// TIA Portal project "Lift" (V15.1)

(* hardware
DEVICE "S7-1200 station_1"  S7-1200 Station
   slot 0: "Rack_0"  S7-1200 Rack  Rack  V1.0
   slot 1: "PLC_1"  CPU 1215C DC/DC/DC  6ES7 215-1AG40-0XB0  V4.2
DEVICE "HMI_1"  TP1500 Basic color PN
   slot 0: "HMI_1"  TP1500 Basic color PN  6AV6 647-0AG11-3AX0  12.0.0.0
   slot 1: "HMI_RT_1"  TP1500 Basic color PN  6AV6 647-0AG11-3AX0  12.0.0.0
   slot 5: "HMI_1.IE_CP_1"  PROFINET Interface  12.0.0.0
      slot 1: "PROFINET Interface_1"  PROFINET Interface
         slot 1: "Port_1"  Port
DEVICE "HMI_2"  KTP700 Basic PN
   slot 0: "HMI_2"  KTP700 Basic PN  6AV2 123-2GB03-0AX0  15.1.0.0
   slot 1: "HMI_RT_2"  KTP700 Basic PN  6AV2 123-2GB03-0AX0  15.1.0.0
   slot 5: "HMI_2.IE_CP_1"  PROFINET Interface  15.0.1.0
      slot 1: "PROFINET Interface_1"  PROFINET Interface
         slot 1: "Port_1"  Port
*)

// ===== PLC "PLC_1"  CPU 1215C DC/DC/DC =====

VAR_GLOBAL   // PLC tag table "Default tag table"
   "Clock_Byte" AT %MB1 : Byte;
   "Clock_10Hz" AT %M1.0 : Bool;
   "Clock_5Hz" AT %M1.1 : Bool;
   "Clock_2.5Hz" AT %M1.2 : Bool;
   "Clock_2Hz" AT %M1.3 : Bool;
   "Clock_1.25Hz" AT %M1.4 : Bool;
   "Clock_1Hz" AT %M1.5 : Bool;
   "Clock_0.625Hz" AT %M1.6 : Bool;
   "Clock_0.5Hz" AT %M1.7 : Bool;
END_VAR

VAR_GLOBAL   // PLC tag table "lift butoane interior"
   "buton_parter" AT %I0.0 : Bool;
   "buton_et1" AT %I0.1 : Bool;
   "buton_et2" AT %I0.2 : Bool;
   "butor_urgenta" AT %I0.3 : Bool;
   "reset_button_urgenta" AT %I0.4 : Bool;
END_VAR

VAR_GLOBAL   // PLC tag table "lift outputs"
   "usa_parter" AT %Q0.0 : Bool;
   "usa_et1" AT %Q0.1 : Bool;
   "usa_et2" AT %Q0.2 : Bool;
   "bec_lift" AT %Q0.3 : Bool;
   "usa lift" AT %Q0.4 : Bool;
END_VAR

VAR_GLOBAL   // PLC tag table "lift auxiliares"
   "block_request_parter" AT %M0.0 : Bool;
   "urgenta_pressed" AT %M2.0 : Bool;
   "block_request_et1" AT %M2.1 : Bool;
   "block_request_et2" AT %M2.2 : Bool;
   "directie sus" AT %M2.3 : Bool;
   "directie jos" AT %M2.4 : Bool;
   "block_persoana" AT %M2.5 : Bool;
   "limitator_parter" AT %M2.6 : Bool;
   "limitator_1" AT %M2.7 : Bool;
   "limitator_2" AT %M3.0 : Bool;
   "reset_block_requests" AT %M3.1 : Bool;
   "tag_auxiliar_hmi" AT %M3.2 : Bool;
END_VAR

VAR_GLOBAL   // PLC tag table "lift butoane exterior"
   "buton_exterior_parter" AT %I0.5 : Bool;
   "buton_et1_ext" AT %I0.6 : Bool;
   "buton_et2_ext" AT %I0.7 : Bool;
END_VAR

VAR_GLOBAL   // PLC tag table "lift inputs(usi)"
   "usa_parter_i" AT %I1.0 : Bool;
   "usa_et1_i" AT %I1.1 : Bool;
   "usa_et2_i" AT %I1.2 : Bool;
   "usa_lift_i" AT %I1.3 : Bool;
END_VAR

DATA_BLOCK "motor_DB"   // DB1
{ S7_Optimized_Access := 'TRUE' }
VERSION : 0.1
// stored: InstanceOfName motor parter
"motor parter"
BEGIN
END_DATA_BLOCK

DATA_BLOCK "motor_DB_1"   // DB2
{ S7_Optimized_Access := 'TRUE' }
VERSION : 0.1
// stored: InstanceOfName motor parter
"motor parter"
BEGIN
END_DATA_BLOCK

DATA_BLOCK "motor_DB_2"   // DB3
{ S7_Optimized_Access := 'TRUE' }
VERSION : 0.1
// stored: InstanceOfName motor parter
"motor parter"
BEGIN
END_DATA_BLOCK

DATA_BLOCK "motor et1_DB"   // DB4
{ S7_Optimized_Access := 'TRUE' }
VERSION : 0.1
// stored: InstanceOfName motor et1
"motor et1"
BEGIN
END_DATA_BLOCK

DATA_BLOCK "motor et2_DB"   // DB5
{ S7_Optimized_Access := 'TRUE' }
VERSION : 0.1
// stored: InstanceOfName motor et2
"motor et2"
BEGIN
END_DATA_BLOCK

DATA_BLOCK "motor parter_DB"   // DB6
{ S7_Optimized_Access := 'TRUE' }
VERSION : 0.1
// stored: InstanceOfName motor parter
"motor parter"
BEGIN
END_DATA_BLOCK

DATA_BLOCK "motor et1_DB_1"   // DB7
{ S7_Optimized_Access := 'TRUE' }
VERSION : 0.1
// stored: InstanceOfName motor et1
"motor et1"
BEGIN
END_DATA_BLOCK

DATA_BLOCK "motor et2_DB_1"   // DB8
{ S7_Optimized_Access := 'TRUE' }
VERSION : 0.1
// stored: InstanceOfName motor et2
"motor et2"
BEGIN
END_DATA_BLOCK

DATA_BLOCK "Commands"   // DB9
{ S7_Optimized_Access := 'TRUE' }
VERSION : 0.1
   VAR
      buton_et1_ext : Bool;
      buton_et2_ext : Bool;
      buton_parter_ext : Bool;
      buton_et1_int : Bool;
      _buton_et2_int : Bool;
      buton_parter_int : Bool;
      buton_urgenta : Bool;
      buton_urgenta_reset : Bool;
      usa_lift_input : Bool;
   END_VAR
BEGIN
END_DATA_BLOCK

FUNCTION_BLOCK "motor parter"   // FB1, LAD
{ S7_Optimized_Access := 'TRUE' }
VERSION : 0.1
   VAR_INPUT
      req_p : Bool;
      et_p : Bool;
      et_1 : Bool;
      et_2 : Bool;
   END_VAR
   VAR_OUTPUT
      dir_sus : Bool;
      dir_jos : Bool;
   END_VAR
BEGIN

REGION Network 1: cerere de la parter
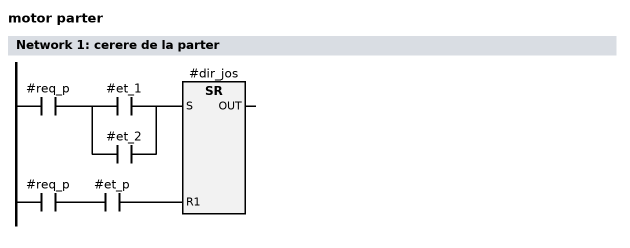
   RUNG wire#powerrail
      Contact( #req_p )
      wire#w1
      Contact( #et_1 )
      wire#w2
      S_SR(operand := #dir_jos, r1 := wire#w3)
   END_RUNG
   RUNG wire#w1
      Contact( #et_2 )
   END_RUNG wire#w2
   RUNG wire#powerrail
      Contact( #req_p )
      Contact( #et_p )
   END_RUNG wire#w3
   // the same network as SCL:
   IF #req_p AND (#et_1 OR #et_2) THEN
       #dir_jos := TRUE;   // SR flip-flop
   END_IF;
   IF #req_p AND #et_p THEN #dir_jos := FALSE; END_IF;
END_REGION
END_FUNCTION_BLOCK

FUNCTION_BLOCK "motor et2"   // FB2, LAD
{ S7_Optimized_Access := 'TRUE' }
VERSION : 0.1
   VAR_INPUT
      req_2 : Bool;
      et_p : Bool;
      et_1 : Bool;
      et_2 : Bool;
   END_VAR
   VAR_OUTPUT
      dir_sus : Bool;
      dir_jos : Bool;
   END_VAR
BEGIN

REGION Network 1: cerere de la etaj 2
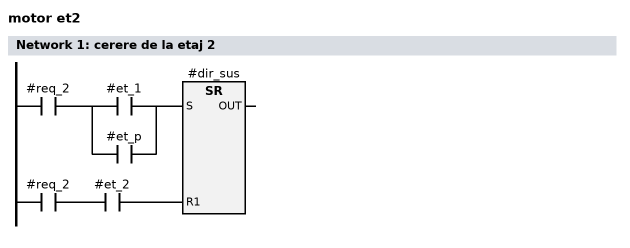
   RUNG wire#powerrail
      Contact( #req_2 )
      wire#w1
      Contact( #et_1 )
      wire#w2
      S_SR(operand := #dir_sus, r1 := wire#w3)
   END_RUNG
   RUNG wire#w1
      Contact( #et_p )
   END_RUNG wire#w2
   RUNG wire#powerrail
      Contact( #req_2 )
      Contact( #et_2 )
   END_RUNG wire#w3
   // the same network as SCL:
   IF #req_2 AND (#et_1 OR #et_p) THEN
       #dir_sus := TRUE;   // SR flip-flop
   END_IF;
   IF #req_2 AND #et_2 THEN #dir_sus := FALSE; END_IF;
END_REGION
END_FUNCTION_BLOCK

FUNCTION_BLOCK "motor et1"   // FB3, LAD
{ S7_Optimized_Access := 'TRUE' }
VERSION : 0.1
   VAR_INPUT
      req_1 : Bool;
      et_p : Bool;
      et_1 : Bool;
      et_2 : Bool;
   END_VAR
   VAR_OUTPUT
      dir_sus : Bool;
      dir_jos : Bool;
   END_VAR
BEGIN

REGION Network 1: cerere de la et 1 venind de la 2
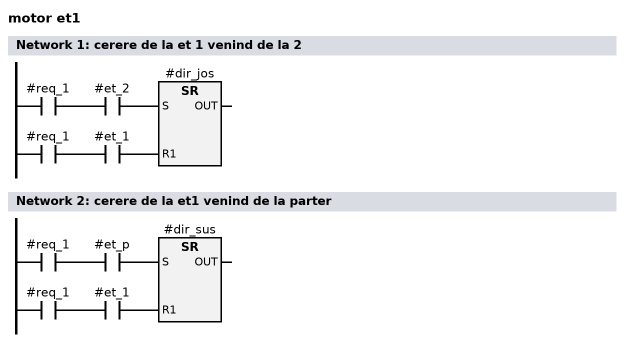
   RUNG wire#powerrail
      Contact( #req_1 )
      Contact( #et_2 )
      S_SR(operand := #dir_jos, r1 := wire#w1)
   END_RUNG
   RUNG wire#powerrail
      Contact( #req_1 )
      Contact( #et_1 )
   END_RUNG wire#w1
   // the same network as SCL:
   IF #req_1 AND #et_2 THEN
       #dir_jos := TRUE;   // SR flip-flop
   END_IF;
   IF #req_1 AND #et_1 THEN #dir_jos := FALSE; END_IF;
END_REGION

REGION Network 2: cerere de la et1 venind de la parter
   RUNG wire#powerrail
      Contact( #req_1 )
      Contact( #et_p )
      S_SR(operand := #dir_sus, r1 := wire#w1)
   END_RUNG
   RUNG wire#powerrail
      Contact( #req_1 )
      Contact( #et_1 )
   END_RUNG wire#w1
   // the same network as SCL:
   IF #req_1 AND #et_p THEN
       #dir_sus := TRUE;   // SR flip-flop
   END_IF;
   IF #req_1 AND #et_1 THEN #dir_sus := FALSE; END_IF;
END_REGION
END_FUNCTION_BLOCK

ORGANIZATION_BLOCK "Main"   // OB1, LAD, ProgramCycle
TITLE = "Main Program Sweep (Cycle)"
{ S7_Optimized_Access := 'TRUE' }
VERSION : 0.1
   VAR_INPUT
      Initial_Call : Bool;   // Initial call of this OB
      Remanence : Bool;   // =True, if remanent data are available
   END_VAR
   VAR_TEMP   // added for the SCL form of the ladder/FBD networks
      _w1 : Bool;
      _w2 : Bool;
      _w3 : Bool;
      _w4 : Bool;
      _w5 : Bool;
      _w6 : Bool;
      _w7 : Bool;
   END_VAR
BEGIN

REGION Network 1: lift butoane pe etaj(sa vina la etajul cerut)
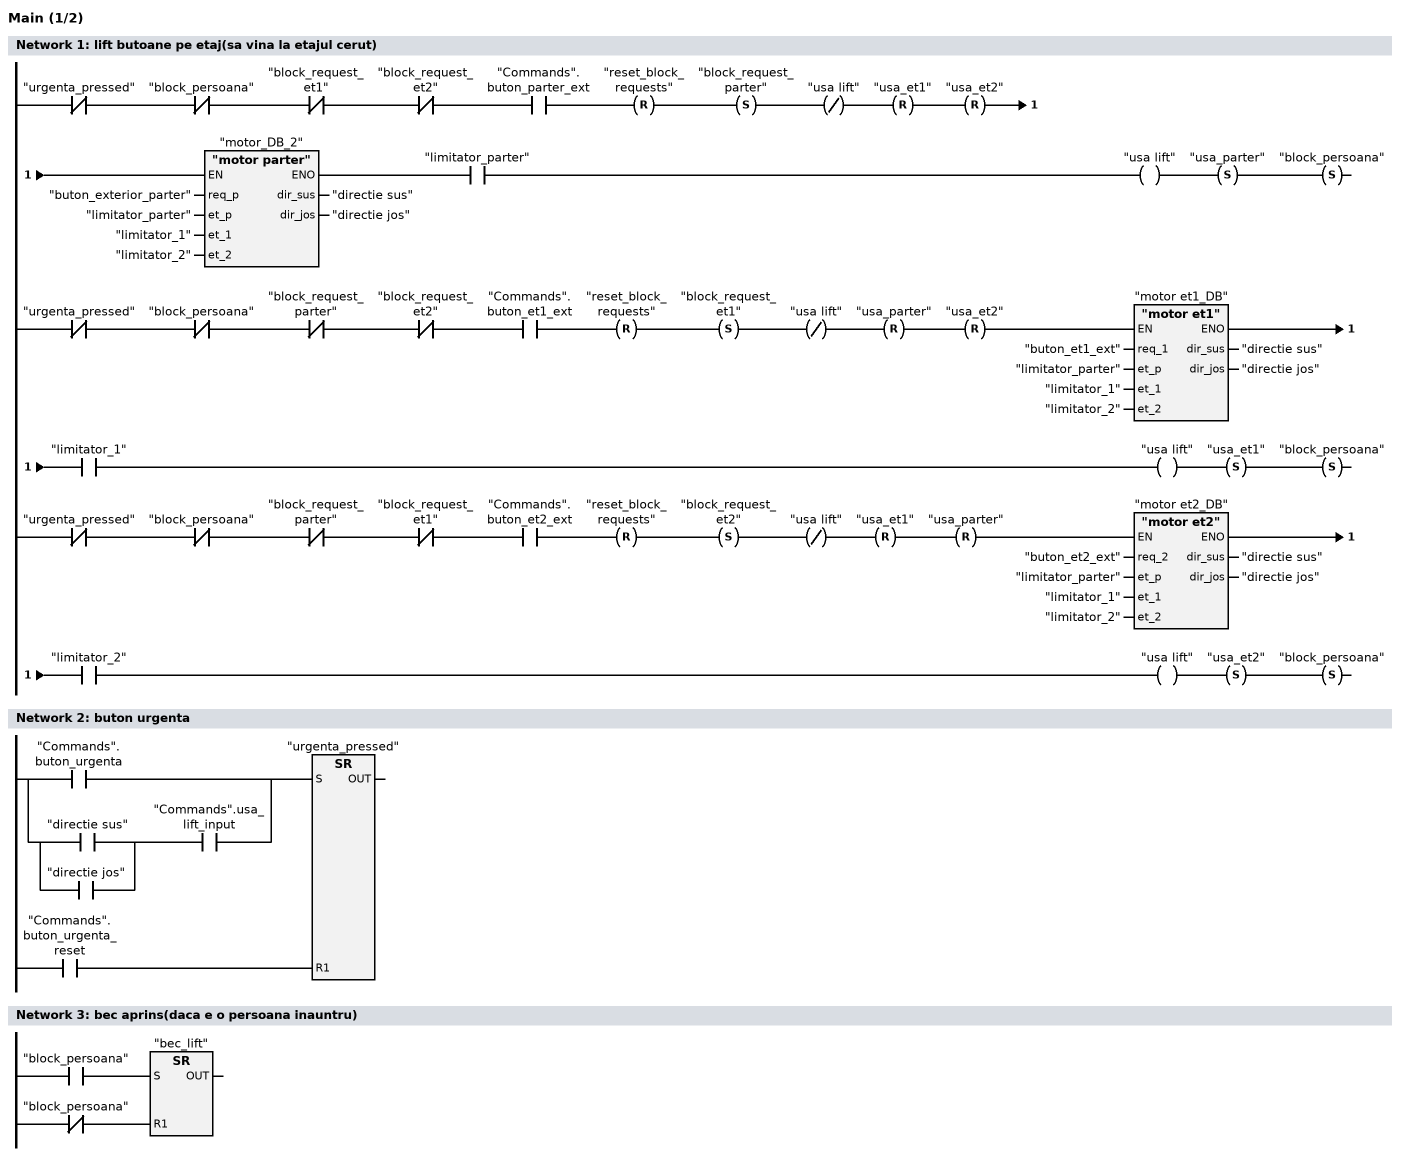
   RUNG wire#powerrail
      I_Contact( "urgenta_pressed" )
      I_Contact( "block_persoana" )
      I_Contact( "block_request_et1" )
      I_Contact( "block_request_et2" )
      Contact( "Commands".buton_parter_ext )
      R_Coil( "reset_block_requests" )
      S_Coil( "block_request_parter" )
      I_Coil( "usa lift" )
      R_Coil( "usa_et1" )
      R_Coil( "usa_et2" )
      "motor_DB_2"(req_p := "buton_exterior_parter", et_p := "limitator_parter", et_1 := "limitator_1", et_2 := "limitator_2", dir_sus => "directie sus", dir_jos => "directie jos")
      Contact( "limitator_parter" )
      Coil( "usa lift" )
      S_Coil( "usa_parter" )
      S_Coil( "block_persoana" )
   END_RUNG
   RUNG wire#powerrail
      I_Contact( "urgenta_pressed" )
      I_Contact( "block_persoana" )
      I_Contact( "block_request_parter" )
      I_Contact( "block_request_et2" )
      Contact( "Commands".buton_et1_ext )
      R_Coil( "reset_block_requests" )
      S_Coil( "block_request_et1" )
      I_Coil( "usa lift" )
      R_Coil( "usa_parter" )
      R_Coil( "usa_et2" )
      "motor et1_DB"(req_1 := "buton_et1_ext", et_p := "limitator_parter", et_1 := "limitator_1", et_2 := "limitator_2", dir_sus => "directie sus", dir_jos => "directie jos")
      Contact( "limitator_1" )
      Coil( "usa lift" )
      S_Coil( "usa_et1" )
      S_Coil( "block_persoana" )
   END_RUNG
   RUNG wire#powerrail
      I_Contact( "urgenta_pressed" )
      I_Contact( "block_persoana" )
      I_Contact( "block_request_parter" )
      I_Contact( "block_request_et1" )
      Contact( "Commands".buton_et2_ext )
      R_Coil( "reset_block_requests" )
      S_Coil( "block_request_et2" )
      I_Coil( "usa lift" )
      R_Coil( "usa_et1" )
      R_Coil( "usa_parter" )
      "motor et2_DB"(req_2 := "buton_et2_ext", et_p := "limitator_parter", et_1 := "limitator_1", et_2 := "limitator_2", dir_sus => "directie sus", dir_jos => "directie jos")
      Contact( "limitator_2" )
      Coil( "usa lift" )
      S_Coil( "usa_et2" )
      S_Coil( "block_persoana" )
   END_RUNG
   // the same network as SCL:
   #_w1 := NOT "urgenta_pressed" AND NOT "block_persoana" AND NOT "block_request_et1" AND NOT "block_request_et2" AND "Commands".buton_parter_ext;
   IF #_w1 THEN
       "reset_block_requests" := FALSE;
       "block_request_parter" := TRUE;
   END_IF;
   "usa lift" := NOT #_w1;
   IF #_w1 THEN
       "usa_et1" := FALSE;
       "usa_et2" := FALSE;
   END_IF;
   "motor_DB_2"(EN := #_w1,   // "motor parter"
                req_p := "buton_exterior_parter",
                et_p := "limitator_parter",
                et_1 := "limitator_1",
                et_2 := "limitator_2",
                dir_sus => "directie sus",
                dir_jos => "directie jos",
                ENO => #_w2);
   "usa lift" := #_w2 AND "limitator_parter";
   IF "usa lift" THEN
       "usa_parter" := TRUE;
       "block_persoana" := TRUE;
   END_IF;
   #_w3 := NOT "urgenta_pressed" AND NOT "block_persoana" AND NOT "block_request_parter" AND NOT "block_request_et2" AND "Commands".buton_et1_ext;
   IF #_w3 THEN
       "reset_block_requests" := FALSE;
       "block_request_et1" := TRUE;
   END_IF;
   "usa lift" := NOT #_w3;
   IF #_w3 THEN
       "usa_parter" := FALSE;
       "usa_et2" := FALSE;
   END_IF;
   "motor et1_DB"(EN := #_w3,   // "motor et1"
                  req_1 := "buton_et1_ext",
                  et_p := "limitator_parter",
                  et_1 := "limitator_1",
                  et_2 := "limitator_2",
                  dir_sus => "directie sus",
                  dir_jos => "directie jos",
                  ENO => #_w4);
   "usa lift" := #_w4 AND "limitator_1";
   IF "usa lift" THEN
       "usa_et1" := TRUE;
       "block_persoana" := TRUE;
   END_IF;
   #_w5 := NOT "urgenta_pressed" AND NOT "block_persoana" AND NOT "block_request_parter" AND NOT "block_request_et1" AND "Commands".buton_et2_ext;
   IF #_w5 THEN
       "reset_block_requests" := FALSE;
       "block_request_et2" := TRUE;
   END_IF;
   "usa lift" := NOT #_w5;
   IF #_w5 THEN
       "usa_et1" := FALSE;
       "usa_parter" := FALSE;
   END_IF;
   "motor et2_DB"(EN := #_w5,   // "motor et2"
                  req_2 := "buton_et2_ext",
                  et_p := "limitator_parter",
                  et_1 := "limitator_1",
                  et_2 := "limitator_2",
                  dir_sus => "directie sus",
                  dir_jos => "directie jos",
                  ENO => #_w6);
   "usa lift" := #_w6 AND "limitator_2";
   IF "usa lift" THEN
       "usa_et2" := TRUE;
       "block_persoana" := TRUE;
   END_IF;
END_REGION

REGION Network 2: buton urgenta
   RUNG wire#powerrail
      Contact( "Commands".buton_urgenta )
      wire#w1
      S_SR(operand := "urgenta_pressed", r1 := wire#w3)
   END_RUNG
   RUNG wire#powerrail
      Contact( "directie sus" )
      wire#w2
      Contact( "Commands".usa_lift_input )
   END_RUNG wire#w1
   RUNG wire#powerrail
      Contact( "directie jos" )
   END_RUNG wire#w2
   RUNG wire#powerrail
      Contact( "Commands".buton_urgenta_reset )
   END_RUNG wire#w3
   // the same network as SCL:
   IF "Commands".buton_urgenta OR (("directie sus" OR "directie jos") AND "Commands".usa_lift_input) THEN
       "urgenta_pressed" := TRUE;   // SR flip-flop
   END_IF;
   IF "Commands".buton_urgenta_reset THEN "urgenta_pressed" := FALSE; END_IF;
END_REGION

REGION Network 3: bec aprins(daca e o persoana inauntru)
   RUNG wire#powerrail
      Contact( "block_persoana" )
      S_SR(operand := "bec_lift", r1 := wire#w1)
   END_RUNG
   RUNG wire#powerrail
      I_Contact( "block_persoana" )
   END_RUNG wire#w1
   // the same network as SCL:
   IF "block_persoana" THEN
       "bec_lift" := TRUE;   // SR flip-flop
   END_IF;
   IF NOT "block_persoana" THEN "bec_lift" := FALSE; END_IF;
END_REGION

REGION Network 4: urcare la etajul cerut
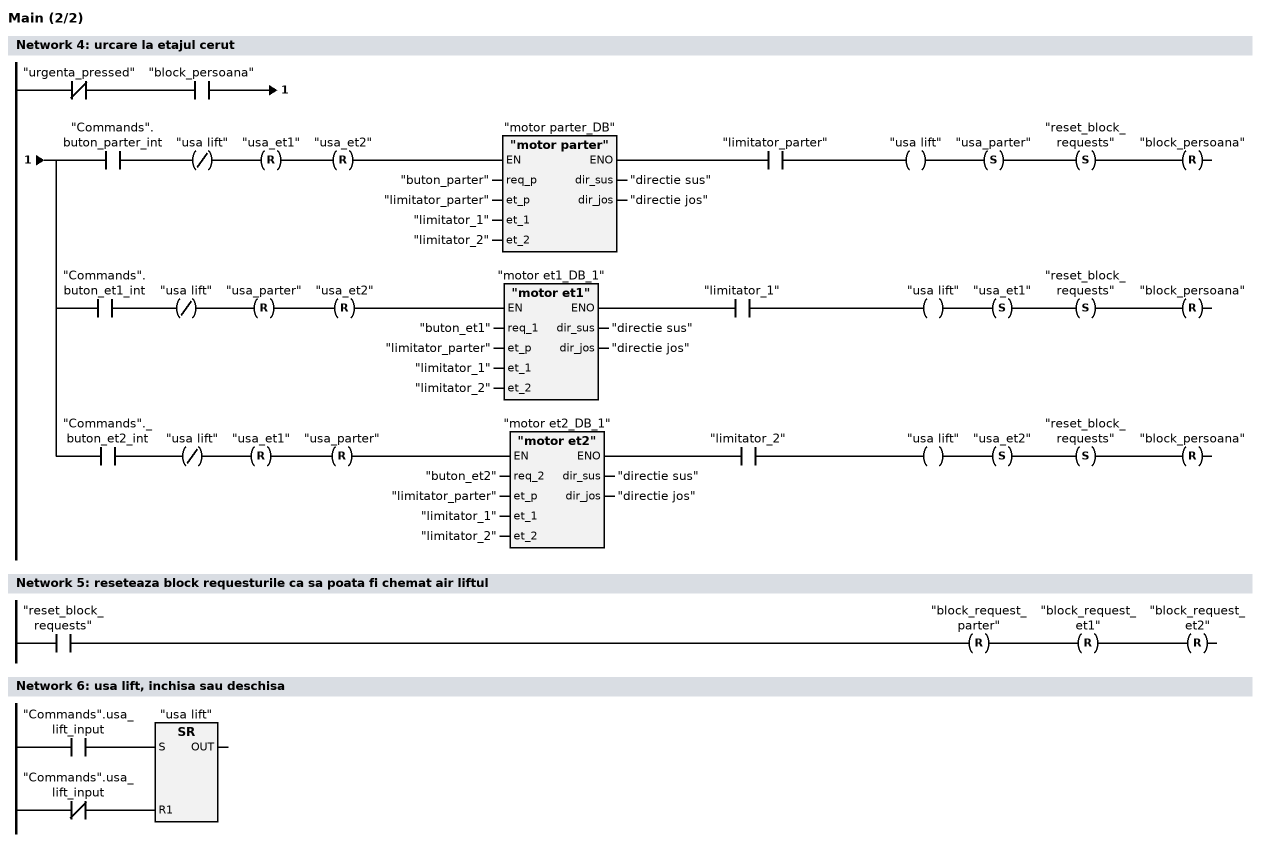
   RUNG wire#powerrail
      I_Contact( "urgenta_pressed" )
      Contact( "block_persoana" )
      wire#w1
      Contact( "Commands".buton_parter_int )
      I_Coil( "usa lift" )
      R_Coil( "usa_et1" )
      R_Coil( "usa_et2" )
      "motor parter_DB"(req_p := "buton_parter", et_p := "limitator_parter", et_1 := "limitator_1", et_2 := "limitator_2", dir_sus => "directie sus", dir_jos => "directie jos")
      Contact( "limitator_parter" )
      Coil( "usa lift" )
      S_Coil( "usa_parter" )
      S_Coil( "reset_block_requests" )
      R_Coil( "block_persoana" )
   END_RUNG
   RUNG wire#w1
      Contact( "Commands".buton_et1_int )
      I_Coil( "usa lift" )
      R_Coil( "usa_parter" )
      R_Coil( "usa_et2" )
      "motor et1_DB_1"(req_1 := "buton_et1", et_p := "limitator_parter", et_1 := "limitator_1", et_2 := "limitator_2", dir_sus => "directie sus", dir_jos => "directie jos")
      Contact( "limitator_1" )
      Coil( "usa lift" )
      S_Coil( "usa_et1" )
      S_Coil( "reset_block_requests" )
      R_Coil( "block_persoana" )
   END_RUNG
   RUNG wire#w1
      Contact( "Commands"._buton_et2_int )
      I_Coil( "usa lift" )
      R_Coil( "usa_et1" )
      R_Coil( "usa_parter" )
      "motor et2_DB_1"(req_2 := "buton_et2", et_p := "limitator_parter", et_1 := "limitator_1", et_2 := "limitator_2", dir_sus => "directie sus", dir_jos => "directie jos")
      Contact( "limitator_2" )
      Coil( "usa lift" )
      S_Coil( "usa_et2" )
      S_Coil( "reset_block_requests" )
      R_Coil( "block_persoana" )
   END_RUNG
   // the same network as SCL:
   #_w1 := NOT "urgenta_pressed" AND "block_persoana";
   #_w2 := #_w1 AND "Commands".buton_parter_int;
   "usa lift" := NOT #_w2;
   IF #_w2 THEN
       "usa_et1" := FALSE;
       "usa_et2" := FALSE;
   END_IF;
   "motor parter_DB"(EN := #_w2,   // "motor parter"
                     req_p := "buton_parter",
                     et_p := "limitator_parter",
                     et_1 := "limitator_1",
                     et_2 := "limitator_2",
                     dir_sus => "directie sus",
                     dir_jos => "directie jos",
                     ENO => #_w3);
   "usa lift" := #_w3 AND "limitator_parter";
   IF "usa lift" THEN
       "usa_parter" := TRUE;
       "reset_block_requests" := TRUE;
       "block_persoana" := FALSE;
   END_IF;
   #_w4 := #_w1 AND "Commands".buton_et1_int;
   "usa lift" := NOT #_w4;
   IF #_w4 THEN
       "usa_parter" := FALSE;
       "usa_et2" := FALSE;
   END_IF;
   "motor et1_DB_1"(EN := #_w4,   // "motor et1"
                    req_1 := "buton_et1",
                    et_p := "limitator_parter",
                    et_1 := "limitator_1",
                    et_2 := "limitator_2",
                    dir_sus => "directie sus",
                    dir_jos => "directie jos",
                    ENO => #_w5);
   "usa lift" := #_w5 AND "limitator_1";
   IF "usa lift" THEN
       "usa_et1" := TRUE;
       "reset_block_requests" := TRUE;
       "block_persoana" := FALSE;
   END_IF;
   #_w6 := #_w1 AND "Commands"._buton_et2_int;
   "usa lift" := NOT #_w6;
   IF #_w6 THEN
       "usa_et1" := FALSE;
       "usa_parter" := FALSE;
   END_IF;
   "motor et2_DB_1"(EN := #_w6,   // "motor et2"
                    req_2 := "buton_et2",
                    et_p := "limitator_parter",
                    et_1 := "limitator_1",
                    et_2 := "limitator_2",
                    dir_sus => "directie sus",
                    dir_jos => "directie jos",
                    ENO => #_w7);
   "usa lift" := #_w7 AND "limitator_2";
   IF "usa lift" THEN
       "usa_et2" := TRUE;
       "reset_block_requests" := TRUE;
       "block_persoana" := FALSE;
   END_IF;
END_REGION

REGION Network 5: reseteaza block requesturile ca sa poata fi chemat air liftul
   RUNG wire#powerrail
      Contact( "reset_block_requests" )
      R_Coil( "block_request_parter" )
      R_Coil( "block_request_et1" )
      R_Coil( "block_request_et2" )
   END_RUNG
   // the same network as SCL:
   IF "reset_block_requests" THEN
       "block_request_parter" := FALSE;
       "block_request_et1" := FALSE;
       "block_request_et2" := FALSE;
   END_IF;
END_REGION

REGION Network 6: usa lift, inchisa sau deschisa
   RUNG wire#powerrail
      Contact( "Commands".usa_lift_input )
      S_SR(operand := "usa lift", r1 := wire#w1)
   END_RUNG
   RUNG wire#powerrail
      I_Contact( "Commands".usa_lift_input )
   END_RUNG wire#w1
   // the same network as SCL:
   IF "Commands".usa_lift_input THEN
       "usa lift" := TRUE;   // SR flip-flop
   END_IF;
   IF NOT "Commands".usa_lift_input THEN "usa lift" := FALSE; END_IF;
END_REGION
END_ORGANIZATION_BLOCK

(* ===== HMI "HMI_RT_1" =====
system functions are stored by id; their names below are inferred from use
connection "HMI_Connection_1": ETHERNET, SMART_S7_1200_OMS

HMI tags "Default tag table"
   "block_persoana" : Bool = PLC block_persoana AT %M2.5, 1 s
   "limitator_1" : Bool = PLC limitator_1 AT %M2.7, 1 s
   "limitator_parter" : Bool = PLC limitator_parter AT %M2.6, 1 s
   "limitator_2" : Bool = PLC limitator_2 AT %M3.0, 1 s
   "Commands_usa_lift_input" : Bool = PLC Commands.usa_lift_input, 1 s
   "Commands_buton_urgenta" : Bool = PLC Commands.buton_urgenta, 1 s
   "Commands_buton_urgenta_reset" : Bool = PLC Commands.buton_urgenta_reset, 1 s
   "Commands_buton_parter_ext" : Bool = PLC Commands.buton_parter_ext, 1 s
   "Commands_buton_et1_ext" : Bool = PLC Commands.buton_et1_ext, 1 s
   "Commands_buton_et2_ext" : Bool = PLC Commands.buton_et2_ext, 1 s
   "Commands_buton_parter_int" : Bool = PLC Commands.buton_parter_int, 1 s
   "Commands_buton_et1_int" : Bool = PLC Commands.buton_et1_int, 1 s
   "Commands__buton_et2_int" : Bool = PLC Commands._buton_et2_int, 1 s
   "Tag_ScreenNumber" : Bool = PLC tag_auxiliar_hmi AT %M3.2, 1 s

Template "Template_1" 1024x768
   Button "Exit" at 943,707 size 79x59; TextOff 'Exit'; PictureOff "ExitRuntime_TP1500_Basic_color_PN"; PictureOn "ExitRuntime_TP1500_Basic_color_PN"
      on Release: StopRuntime(0)
   Button "Template_Button" at 857,707 size 79x59; TextOff 'Text'
   Button "Template_Button_1" at 772,707 size 79x59; TextOff 'Text'
   Button "Template_Button_2" at 686,707 size 79x59; TextOff 'Text'
   Button "Template_Button_3" at 600,707 size 79x59; TextOff 'Text'
   Button "Template_Button_4" at 515,707 size 79x59; TextOff 'Text'
   Button "Template_Button_5" at 429,707 size 79x59; TextOff 'Text'
   Button "Template_Button_6" at 344,707 size 79x59; TextOff 'Text'
   Button "Template_Button_7" at 258,707 size 79x59; TextOff 'Text'
   Button "Template_Button_8" at 172,707 size 79x59; TextOff 'Text'
   Button "Alarms" at 87,707 size 79x59; TextOff 'Alarms'; PictureOff "AlarmDisplay_TP1500_Basic_color_PN"; PictureOn "AlarmDisplay_TP1500_Basic_color_PN"
      on Release: function_ef3f5d25("Alarm window_Unacknowledged", -1)
   Button "Start screen" at 1,707 size 79x59; TextOff 'Start screen'; PictureOff "NavigateHome_TP1500_Basic_color_PN"; PictureOn "NavigateHome_TP1500_Basic_color_PN"
      on Release: ActivateScreen("Root screen", 0)
   DateTimeField "HmiScreenItemData" at 919,30 size 105x30
   DateTimeField "HmiScreenItemData_1" at 919,0 size 105x30

screen "Root screen" 1024x768, template "Template_1"
   Rectangle "Rectangle_1" at 324,269 size 72x35
      Appearance <- "limitator_parter"
   Rectangle "Rectangle_2" at 324,212 size 72x35
      Appearance <- "limitator_1"
   Rectangle "Rectangle_3" at 324,150 size 72x35
      Appearance <- "limitator_2"
   TextField "Text field_1" at 262,280 size 50x20; Text 'Parter'
   TextField "Text field_2" at 261,227 size 27x20; Text 'Et1'
   TextField "Text field_3" at 268,166 size 27x20; Text 'Et2'
   TextField "Text field_4" at 731,70 size 63x20; Text 'Exterior'
   TextField "Text field_5" at 878,70 size 61x20; Text 'Interior'
   Button "Button_7" at 422,76 size 72x23; TextOff 'Urgenta'
      on Click: SetBit("Commands_buton_urgenta")
   Button "Button_8" at 519,76 size 72x23; TextOff 'Reset Urg'
      on Click: SetBit("Commands_buton_urgenta_reset")
   Circle "Circle_1" at 520,204 size 61x61
      Appearance <- "block_persoana"
   TextField "Text field_6" at 520,186 size 72x20; Text 'Persoana'
   Button "Button_9" at 781,288 size 72x23; TextOff 'Inchide'
      on Click: ResetBit("Commands_usa_lift_input")
   Button "Button_10" at 878,288 size 72x23; TextOff 'Deschide'
      on Click: SetBit("Commands_usa_lift_input")
   TextField "Text field_7" at 834,259 size 96x20; Text 'Usa de la lift'
   TextField "Text field_8" at 467,338 size 83x20; Text 'A ajuns la:'
   Button "Button_14" at 649,26 size 72x23; TextOff 'Reset'
   Switch "Switch_1" at 467,363 size 57x23; CaptionText 'Switch'; TextOff 'OFF'; TextOn 'ON'
      on SwitchOn: SetBit("limitator_parter"); ResetBit("limitator_1"); ResetBit("limitator_2")
      on SwitchOff: ResetBit("limitator_parter")
   TextField "Text field_9" at 479,406 size 50x20; Text 'Parter'
   TextField "Text field_10" at 721,406 size 12x20; Text '2'
   TextField "Text field_11" at 590,398 size 12x20; Text '1'
   Switch "Switch_2" at 574,363 size 57x23; TextOn 'ON'; CaptionText 'Switch'; TextOff 'OFF'
      on SwitchOff: ResetBit("limitator_1")
      on SwitchOn: SetBit("limitator_1"); ResetBit("limitator_parter"); ResetBit("limitator_2")
   Switch "Switch_3" at 698,363 size 57x23; TextOn 'ON'; CaptionText 'Switch'; TextOff 'OFF'
      on SwitchOff: ResetBit("limitator_2")
      on SwitchOn: SetBit("limitator_2"); ResetBit("limitator_1"); ResetBit("limitator_parter")
   TextField "Text field_12" at 668,104 size 50x20; Text 'Parter'
   TextField "Text field_13" at 683,147 size 12x20; Text '1'
   TextField "Text field_14" at 684,189 size 12x20; Text '2'
   Switch "Switch_4" at 740,104 size 57x23; TextOn 'ON'; CaptionText 'Switch'; TextOff 'OFF'
      on SwitchOff: ResetBit("Commands_buton_parter_ext")
      on SwitchOn: SetBit("Commands_buton_parter_ext")
   Switch "Switch_5" at 860,143 size 57x23; TextOn 'ON'; CaptionText 'Switch'; TextOff 'OFF'
      on SwitchOn: SetBit("Commands_buton_et1_int")
      on SwitchOff: ResetBit("Commands_buton_et1_int")
   Switch "Switch_6" at 860,104 size 57x23; TextOn 'ON'; CaptionText 'Switch'; TextOff 'OFF'
      on SwitchOn: SetBit("Commands_buton_parter_int")
      on SwitchOff: ResetBit("Commands_buton_parter_int")
   Switch "Switch_7" at 741,180 size 57x23; TextOn 'ON'; CaptionText 'Switch'; TextOff 'OFF'
      on SwitchOn: SetBit("Commands_buton_et2_ext")
      on SwitchOff: ResetBit("Commands_buton_et2_ext")
   Switch "Switch_8" at 740,143 size 57x23; TextOn 'ON'; CaptionText 'Switch'; TextOff 'OFF'
      on SwitchOn: SetBit("Commands_buton_et1_ext")
      on SwitchOff: ResetBit("Commands_buton_et1_ext")
   Switch "Switch_9" at 860,181 size 57x23; TextOn 'ON'; CaptionText 'Switch'; TextOff 'OFF'
      on SwitchOn: SetBit("Commands__buton_et2_int")
      on SwitchOff: ResetBit("Commands__buton_et2_int")
   Button "Button_1" at 310,363 size 72x23; TextOff 'Parter'
      on Click: SetBit("limitator_parter"); ResetBit("limitator_1"); ResetBit("limitator_2")
   Button "Button_2" at 297,394 size 72x23; TextOff 'Etaj 1'
      on Click: SetBit("limitator_1"); ResetBit("limitator_parter"); ResetBit("limitator_2")
   Button "Button_3" at 283,426 size 72x23; TextOff 'Etaj 2'
      on Click: SetBit("limitator_2"); ResetBit("limitator_1"); ResetBit("limitator_parter")
   Group "Group" at 261,26 size 689x423

screen "Screen_1" 1024x768
   AlarmView "Alarm view_1" at 0,0 size 1023x767
*)

(* ===== HMI "HMI_RT_2" =====
system functions are stored by id; their names below are inferred from use
connection "HMI_Connection_2": ETHERNET, SMART_S7_1200_OMS

HMI tags "Default tag table"
   "Tag_ScreenNumber" : UInt, internal
   "motor et2_DB_req_2" : Bool = PLC "motor et2_DB".req_2, 1 s
   "block_persoana" : Bool = PLC block_persoana AT %M2.5, 1 s
   "Commands__buton_et2_int" : Bool = PLC Commands._buton_et2_int, 1 s
   "Commands_buton_et1_ext" : Bool = PLC Commands.buton_et1_ext, 1 s
   "Commands_buton_et1_int" : Bool = PLC Commands.buton_et1_int, 1 s
   "Commands_buton_et2_ext" : Bool = PLC Commands.buton_et2_ext, 1 s
   "Commands_buton_parter_ext" : Bool = PLC Commands.buton_parter_ext, 1 s
   "Commands_buton_parter_int" : Bool = PLC Commands.buton_parter_int, 1 s
   "Commands_buton_urgenta" : Bool = PLC Commands.buton_urgenta, 1 s
   "Commands_buton_urgenta_reset" : Bool = PLC Commands.buton_urgenta_reset, 1 s
   "Commands_usa_lift_input" : Bool = PLC Commands.usa_lift_input, 1 s
   "limitator_1" : Bool = PLC limitator_1 AT %M2.7, 1 s
   "limitator_2" : Bool = PLC limitator_2 AT %M3.0, 1 s
   "limitator_parter" : Bool = PLC limitator_parter AT %M2.6, 1 s
   "Tag_ScreenNumber(1)" : Bool = PLC tag_auxiliar_hmi AT %M3.2, 1 s

Template "Template_1" 800x480
   Button "Exit" at 714,429 size 71x50; TextOff 'Exit'; PictureOff "ExitRuntime_KTP700_Basic_PN_TR"; PictureOn "ExitRuntime_KTP700_Basic_PN_TR"
      on Release: StopRuntime(0)
   Button "Template_Button" at 614,429 size 71x50; TextOff 'Text'
   Button "Template_Button_1" at 514,429 size 71x50; TextOff 'Text'
   Button "Template_Button_2" at 414,429 size 71x50; TextOff 'Text'
   Button "Template_Button_3" at 314,429 size 71x50; TextOff 'Text'
   Button "Template_Button_4" at 214,429 size 71x50; TextOff 'Text'
   Button "Template_Button_5" at 114,429 size 71x50; TextOff 'Text'
   Button "Start screen" at 14,429 size 71x50; TextOff 'Start screen'; PictureOff "NavigateHome_KTP700_Basic_PN_TR"; PictureOn "NavigateHome_KTP700_Basic_PN_TR"
      on Release: ActivateScreen("Root screen", 0)
   SymbolicIOField "Symbolic_IO_Field_Screen" at 93,9 size 600x33; TextOff '0'; TextOn '1'; TextList "TextList_ScreenNames"
      ProcessValue <- "Tag_ScreenNumber"
      on Change: ActivateScreenByNumber("Tag_ScreenNumber", 0)
   DateTimeField "HmiScreenItemData" at 695,25 size 105x25
   DateTimeField "HmiScreenItemData_1" at 695,0 size 105x25
   GraphicView "Logo" at 0,0 size 91x51; Picture "Logo of HMI_2"

screen "Root screen" 800x480, template "Template_1"
   on GenerateScreen: SetTag("Tag_ScreenNumber", 1)
   Rectangle "Rectangle_1" at 90,261 size 76x30
      Appearance <- "limitator_parter"
   Rectangle "Rectangle_2" at 90,212 size 76x30
      Appearance <- "limitator_1"
   Rectangle "Rectangle_3" at 90,159 size 76x30
      Appearance <- "limitator_2"
   TextField "Text field_1" at 25,270 size 50x20; Text 'Parter'
   TextField "Text field_2" at 23,225 size 27x20; Text 'Et1'
   TextField "Text field_3" at 31,172 size 27x20; Text 'Et2'
   TextField "Text field_4" at 523,90 size 63x20; Text 'Exterior'
   TextField "Text field_5" at 680,90 size 61x20; Text 'Interior'
   Circle "Circle_1" at 305,208 size 53x53
      Appearance <- "block_persoana"
   TextField "Text field_6" at 299,190 size 72x20; Text 'Persoana'
   Button "Button_9" at 576,278 size 76x20; TextOff 'Inchide'
      on Click: ResetBit("Commands_usa_lift_input")
   Button "Button_10" at 680,278 size 76x20; TextOff 'Deschide'
      on Click: SetBit("Commands_usa_lift_input")
   TextField "Text field_7" at 632,253 size 96x20; Text 'Usa de la lift'
   TextField "Text field_8" at 242,321 size 83x20; Text 'A ajuns la:'
   Button "Button_14" at 436,52 size 76x20; TextOff 'Reset'
   Switch "Switch_1" at 242,342 size 61x20; TextOn 'ON'; CaptionText 'Switch'; TextOff 'OFF'
      on SwitchOff: ResetBit("limitator_parter")
      on SwitchOn: SetBit("limitator_parter"); ResetBit("limitator_1"); ResetBit("limitator_2")
   TextField "Text field_9" at 255,379 size 50x20; Text 'Parter'
   TextField "Text field_10" at 512,379 size 12x20; Text '2'
   TextField "Text field_11" at 373,372 size 12x20; Text '1'
   Switch "Switch_2" at 356,342 size 61x20; TextOn 'ON'; CaptionText 'Switch'; TextOff 'OFF'
      on SwitchOn: SetBit("limitator_1"); ResetBit("limitator_parter"); ResetBit("limitator_2")
      on SwitchOff: ResetBit("limitator_1")
   Switch "Switch_3" at 488,342 size 61x20; TextOn 'ON'; CaptionText 'Switch'; TextOff 'OFF'
      on SwitchOn: SetBit("limitator_2"); ResetBit("limitator_1"); ResetBit("limitator_parter")
      on SwitchOff: ResetBit("limitator_2")
   TextField "Text field_12" at 456,119 size 50x20; Text 'Parter'
   TextField "Text field_13" at 472,156 size 12x20; Text '1'
   TextField "Text field_14" at 473,192 size 12x20; Text '2'
   Switch "Switch_4" at 533,119 size 61x20; TextOn 'ON'; CaptionText 'Switch'; TextOff 'OFF'
      on SwitchOn: SetBit("Commands_buton_parter_ext")
      on SwitchOff: ResetBit("Commands_buton_parter_ext")
   Switch "Switch_5" at 661,152 size 61x20; TextOn 'ON'; CaptionText 'Switch'; TextOff 'OFF'
      on SwitchOff: ResetBit("Commands_buton_et1_int")
      on SwitchOn: SetBit("Commands_buton_et1_int")
   Switch "Switch_6" at 661,119 size 61x20; TextOn 'ON'; CaptionText 'Switch'; TextOff 'OFF'
      on SwitchOff: ResetBit("Commands_buton_parter_int")
      on SwitchOn: SetBit("Commands_buton_parter_int")
   Switch "Switch_7" at 534,185 size 61x20; TextOn 'ON'; CaptionText 'Switch'; TextOff 'OFF'
      on SwitchOff: ResetBit("Commands_buton_et2_ext")
      on SwitchOn: SetBit("Commands_buton_et2_ext")
   Switch "Switch_8" at 533,152 size 61x20; TextOn 'ON'; CaptionText 'Switch'; TextOff 'OFF'
      on SwitchOff: ResetBit("Commands_buton_et1_ext")
      on SwitchOn: SetBit("Commands_buton_et1_ext")
   Switch "Switch_9" at 661,185 size 61x20; TextOn 'ON'; CaptionText 'Switch'; TextOff 'OFF'
      on SwitchOff: ResetBit("Commands__buton_et2_int")
      on SwitchOn: SetBit("Commands__buton_et2_int")
   Switch "Switch_10" at 203,119 size 61x20; TextOn 'ON'; CaptionText 'Switch'; TextOff 'OFF'
      on SwitchOff: ResetBit("Commands_buton_urgenta")
      on SwitchOn: SetBit("Commands_buton_urgenta")
   Switch "Switch_11" at 303,124 size 61x20; TextOn 'ON'; CaptionText 'Switch'; TextOff 'OFF'
      on SwitchOff: ResetBit("Commands_buton_urgenta_reset")
      on SwitchOn: SetBit("Commands_buton_urgenta_reset")
   TextField "Text field_15" at 189,91 size 71x23; Text 'Urgenta'
   TextField "Text field_16" at 290,91 size 123x23; Text 'Reset Urgenta'
*)